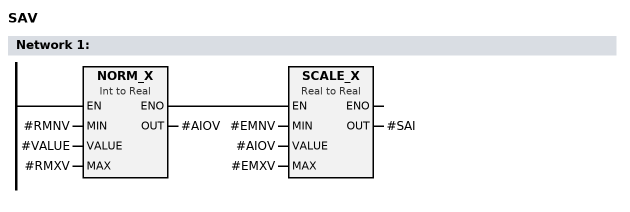
   RUNG wire#powerrail
      { S7_Templates := "[SrcType := Int, DestType := Real]" } Normalize(min := #RMNV, value := #VALUE, max := #RMXV, out => #AIOV)
      { S7_Templates := "[SrcType := Real, DestType := Real]" } Scale(min := #EMNV, value := #AIOV, max := #EMXV, out => #SAI)
   END_RUNG
   // the same network as SCL:
   #AIOV := NORM_X(MIN := #RMNV, VALUE := #VALUE, MAX := #RMXV);
   #SAI := SCALE_X(MIN := #EMNV, VALUE := #AIOV, MAX := #EMXV);
END_REGION
END_FUNCTION

// folder: 1}Library/Interlock

FUNCTION_BLOCK "Interlocks"   // FB4550, LAD
{ S7_Optimized_Access := 'TRUE' }
VERSION : 0.1
   VAR_INPUT
      Interlock_1 : Bool;
      Interlock_2 : Bool;
      Interlock_3 : Bool;
      Interlock_4 : Bool;
      Interlock_5 : Bool := false;
      Interlock_6 : Bool := false;
      Interlock_7 : Bool := false;
      Interlock_8 : Bool := false;
      Interlock_9 : Bool := false;
      Interlock_10 : Bool := false;
      Interlock_11 : Bool := false;
      Interlock_12 : Bool := false;
      Interlock_13 : Bool := false;
      Interlock_14 : Bool := false;
      Interlock_15 : Bool := false;
      Interlock_16 : Bool := false;
      Interlock_17 : Bool := false;
      Interlock_18 : Bool := false;
      Interlock_19 : Bool := false;
      Interlock_20 : Bool := false;
      Interlock_21 : Bool := false;
      Interlock_22 : Bool := false;
      Interlock_23 : Bool := false;
      Interlock_24 : Bool := false;
      Interlock_25 : Bool := false;
      Interlock_26 : Bool := false;
      Interlock_27 : Bool := false;
      Interlock_28 : Bool := false;
      Interlock_29 : Bool := false;
      Interlock_30 : Bool := false;
      Interlock_31 : Bool := false;
      Interlock_32 : Bool := false;
   END_VAR
   VAR_OUTPUT
      Out : Bool;   // Common Interlock Output
      Latched_Interlocks : DInt;   // Status of all Interlocks
   END_VAR
   VAR_IN_OUT
      Reset : Bool;
   END_VAR
   VAR
      HMI : Struct
         Interlock_1 : Bool;
         Interlock_2 : Bool;
         Interlock_3 : Bool;
         Interlock_4 : Bool;
         Interlock_5 : Bool;
         Interlock_6 : Bool;
         Interlock_7 : Bool;
         Interlock_8 : Bool;
         Interlock_9 : Bool;
         Interlock_10 : Bool;
         Interlock_11 : Bool;
         Interlock_12 : Bool;
         Interlock_13 : Bool;
         Interlock_14 : Bool;
         Interlock_15 : Bool;
         Interlock_16 : Bool;
         Interlock_17 : Bool;
         Interlock_18 : Bool;
         Interlock_19 : Bool;
         Interlock_20 : Bool;
         Interlock_21 : Bool;
         Interlock_22 : Bool;
         Interlock_23 : Bool;
         Interlock_24 : Bool;
         Interlock_25 : Bool;
         Interlock_26 : Bool;
         Interlock_27 : Bool;
         Interlock_28 : Bool;
         Interlock_29 : Bool;
         Interlock_30 : Bool;
         Interlock_31 : Bool;
         Interlock_32 : Bool;
         First_1 : Bool;
         First_2 : Bool;
         First_3 : Bool;
         First_4 : Bool;
         First_5 : Bool;
         First_6 : Bool;
         First_7 : Bool;
         First_8 : Bool;
         First_9 : Bool;
         First_10 : Bool;
         First_11 : Bool;
         First_12 : Bool;
         First_13 : Bool;
         First_14 : Bool;
         First_15 : Bool;
         First_16 : Bool;
         First_17 : Bool;
         First_18 : Bool;
         First_19 : Bool;
         First_20 : Bool;
         First_21 : Bool;
         First_22 : Bool;
         First_23 : Bool;
         First_24 : Bool;
         First_25 : Bool;
         First_26 : Bool;
         First_27 : Bool;
         First_28 : Bool;
         First_29 : Bool;
         First_30 : Bool;
         First_31 : Bool;
         First_32 : Bool;
         Bypass_1 : Bool;
         Bypass_2 : Bool;
         Bypass_3 : Bool;
         Bypass_4 : Bool;
         Bypass_5 : Bool;
         Bypass_6 : Bool;
         Bypass_7 : Bool;
         Bypass_8 : Bool;
         Bypass_9 : Bool;
         Bypass_10 : Bool;
         Bypass_11 : Bool;
         Bypass_12 : Bool;
         Bypass_13 : Bool;
         Bypass_14 : Bool;
         Bypass_15 : Bool;
         Bypass_16 : Bool;
         Bypass_17 : Bool;
         Bypass_18 : Bool;
         Bypass_19 : Bool;
         Bypass_20 : Bool;
         Bypass_21 : Bool;
         Bypass_22 : Bool;
         Bypass_23 : Bool;
         Bypass_24 : Bool;
         Bypass_25 : Bool;
         Bypass_26 : Bool;
         Bypass_27 : Bool;
         Bypass_28 : Bool;
         Bypass_29 : Bool;
         Bypass_30 : Bool;
         Bypass_31 : Bool;
         Bypass_32 : Bool;
         Status_DW : DInt;
         Interlock_DW : DInt;
         First_DW : DInt;
         Bypass_DW : DInt;
      END_STRUCT;
   END_VAR
   VAR_TEMP
      Initial_Trip : Bool;
      Interlocks_Status : DInt;
   END_VAR
BEGIN

REGION Network 1 (SCL): Common Interlock Input
   ;
   #Interlocks_Status.%X0:= #Interlock_1;
   #Interlocks_Status.%X1 := #Interlock_2;
   #Interlocks_Status.%X2 := #Interlock_3;
   #Interlocks_Status.%X3 := #Interlock_4;
   #Interlocks_Status.%X4 := #Interlock_5;
   #Interlocks_Status.%X5 := #Interlock_6;
   #Interlocks_Status.%X6 := #Interlock_7;
   #Interlocks_Status.%X7 := #Interlock_8;
   #Interlocks_Status.%X8 := #Interlock_9;
   #Interlocks_Status.%X9 := #Interlock_10;
   #Interlocks_Status.%X10 := #Interlock_11;
   #Interlocks_Status.%X11 := #Interlock_12;
   #Interlocks_Status.%X12 := #Interlock_13;
   #Interlocks_Status.%X13 := #Interlock_14;
   #Interlocks_Status.%X14 := #Interlock_15;
   #Interlocks_Status.%X15 := #Interlock_16;
   #Interlocks_Status.%X16 := #Interlock_17;
   #Interlocks_Status.%X17 := #Interlock_18;
   #Interlocks_Status.%X18 := #Interlock_19;
   #Interlocks_Status.%X19 := #Interlock_20;
   #Interlocks_Status.%X20 := #Interlock_21;
   #Interlocks_Status.%X21 := #Interlock_22;
   #Interlocks_Status.%X22 := #Interlock_23;
   #Interlocks_Status.%X23 := #Interlock_24;
   #Interlocks_Status.%X24 := #Interlock_25;
   #Interlocks_Status.%X25 := #Interlock_26;
   #Interlocks_Status.%X26 := #Interlock_27;
   #Interlocks_Status.%X27 := #Interlock_28;
   #Interlocks_Status.%X28 := #Interlock_29;
   #Interlocks_Status.%X29 := #Interlock_30;
   #Interlocks_Status.%X30 := #Interlock_31;
   #Interlocks_Status.%X31 := #Interlock_32;
END_REGION

REGION Network 2 (SCL): Bypass Move
   #HMI.Bypass_1 := #HMI.Bypass_DW.%X0;
   #HMI.Bypass_2 := #HMI.Bypass_DW.%X1;
   #HMI.Bypass_3 := #HMI.Bypass_DW.%X2;
   #HMI.Bypass_4 := #HMI.Bypass_DW.%X3;
   #HMI.Bypass_5 := #HMI.Bypass_DW.%X4;
   #HMI.Bypass_6 := #HMI.Bypass_DW.%X5;
   #HMI.Bypass_7 := #HMI.Bypass_DW.%X6;
   #HMI.Bypass_8 := #HMI.Bypass_DW.%X7;
   #HMI.Bypass_9 := #HMI.Bypass_DW.%X8;
   #HMI.Bypass_10 := #HMI.Bypass_DW.%X9;
   #HMI.Bypass_11 := #HMI.Bypass_DW.%X10;
   #HMI.Bypass_12 := #HMI.Bypass_DW.%X11;
   #HMI.Bypass_13 := #HMI.Bypass_DW.%X12;
   #HMI.Bypass_14 := #HMI.Bypass_DW.%X13;
   #HMI.Bypass_15 := #HMI.Bypass_DW.%X14;
   #HMI.Bypass_16 := #HMI.Bypass_DW.%X15;
   #HMI.Bypass_17 := #HMI.Bypass_DW.%X16;
   #HMI.Bypass_18 := #HMI.Bypass_DW.%X17;
   #HMI.Bypass_19 := #HMI.Bypass_DW.%X18;
   #HMI.Bypass_20 := #HMI.Bypass_DW.%X19;
   #HMI.Bypass_21 := #HMI.Bypass_DW.%X20;
   #HMI.Bypass_22 := #HMI.Bypass_DW.%X21;
   #HMI.Bypass_23 := #HMI.Bypass_DW.%X22;
   #HMI.Bypass_24 := #HMI.Bypass_DW.%X23;
   #HMI.Bypass_25 := #HMI.Bypass_DW.%X24;
   #HMI.Bypass_26 := #HMI.Bypass_DW.%X25;
   #HMI.Bypass_27 := #HMI.Bypass_DW.%X26;
   #HMI.Bypass_28 := #HMI.Bypass_DW.%X27;
   #HMI.Bypass_29 := #HMI.Bypass_DW.%X28;
   #HMI.Bypass_30 := #HMI.Bypass_DW.%X29;
   #HMI.Bypass_31 := #HMI.Bypass_DW.%X30;
   #HMI.Bypass_32 := #HMI.Bypass_DW.%X31;
END_REGION

REGION Network 3: Match HMI.Status_DW to Interlocks_Status
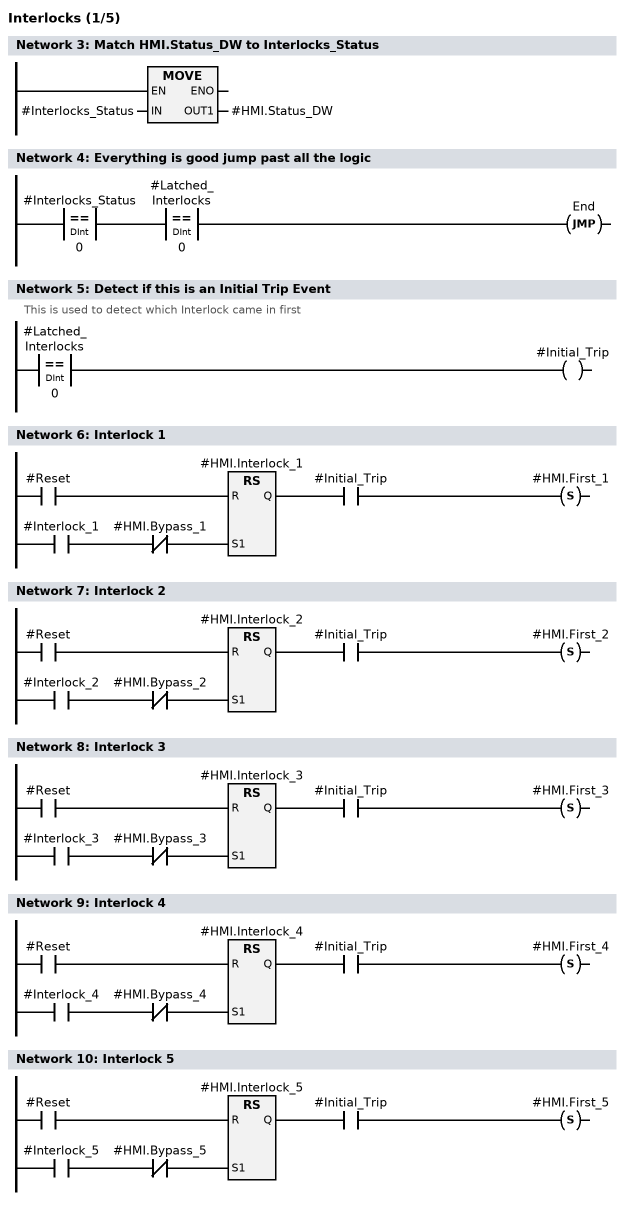
   RUNG wire#powerrail
      Move(in := #Interlocks_Status, out1 => #HMI.Status_DW)
   END_RUNG
   // the same network as SCL:
   #HMI.Status_DW := #Interlocks_Status;
END_REGION

REGION Network 4: Everything is good jump past all the logic
   RUNG wire#powerrail
      { S7_Templates := "SrcType := DInt" } EQ_Contact(in1 := #Interlocks_Status, in2 := 0)
      { S7_Templates := "SrcType := DInt" } EQ_Contact(in1 := #Latched_Interlocks, in2 := 0)
      JumpCoil( End )
   END_RUNG
   // the same network as SCL:
   IF (#Interlocks_Status = 0) AND (#Latched_Interlocks = 0) THEN GOTO End; END_IF;
END_REGION

REGION Network 5: Detect if this is an Initial Trip Event
   // This is used to detect which Interlock came in first
   RUNG wire#powerrail
      { S7_Templates := "SrcType := DInt" } EQ_Contact(in1 := #Latched_Interlocks, in2 := 0)
      Coil( #Initial_Trip )
   END_RUNG
   // the same network as SCL:
   #Initial_Trip := #Latched_Interlocks = 0;
END_REGION

REGION Network 6: Interlock 1
   RUNG wire#powerrail
      Contact( #Reset )
      S_RS(operand := #HMI.Interlock_1, s1 := wire#w1)
      Contact( #Initial_Trip )
      S_Coil( #HMI.First_1 )
   END_RUNG
   RUNG wire#powerrail
      Contact( #Interlock_1 )
      I_Contact( #HMI.Bypass_1 )
   END_RUNG wire#w1
   // the same network as SCL:
   IF #Reset THEN
       #HMI.Interlock_1 := FALSE;   // RS flip-flop
   END_IF;
   IF #Interlock_1 AND NOT #HMI.Bypass_1 THEN #HMI.Interlock_1 := TRUE; END_IF;
   IF #HMI.Interlock_1 AND #Initial_Trip THEN #HMI.First_1 := TRUE; END_IF;
END_REGION

REGION Network 7: Interlock 2
   RUNG wire#powerrail
      Contact( #Reset )
      S_RS(operand := #HMI.Interlock_2, s1 := wire#w1)
      Contact( #Initial_Trip )
      S_Coil( #HMI.First_2 )
   END_RUNG
   RUNG wire#powerrail
      Contact( #Interlock_2 )
      I_Contact( #HMI.Bypass_2 )
   END_RUNG wire#w1
   // the same network as SCL:
   IF #Reset THEN
       #HMI.Interlock_2 := FALSE;   // RS flip-flop
   END_IF;
   IF #Interlock_2 AND NOT #HMI.Bypass_2 THEN #HMI.Interlock_2 := TRUE; END_IF;
   IF #HMI.Interlock_2 AND #Initial_Trip THEN #HMI.First_2 := TRUE; END_IF;
END_REGION

REGION Network 8: Interlock 3
   RUNG wire#powerrail
      Contact( #Reset )
      S_RS(operand := #HMI.Interlock_3, s1 := wire#w1)
      Contact( #Initial_Trip )
      S_Coil( #HMI.First_3 )
   END_RUNG
   RUNG wire#powerrail
      Contact( #Interlock_3 )
      I_Contact( #HMI.Bypass_3 )
   END_RUNG wire#w1
   // the same network as SCL:
   IF #Reset THEN
       #HMI.Interlock_3 := FALSE;   // RS flip-flop
   END_IF;
   IF #Interlock_3 AND NOT #HMI.Bypass_3 THEN #HMI.Interlock_3 := TRUE; END_IF;
   IF #HMI.Interlock_3 AND #Initial_Trip THEN #HMI.First_3 := TRUE; END_IF;
END_REGION

REGION Network 9: Interlock 4
   RUNG wire#powerrail
      Contact( #Reset )
      S_RS(operand := #HMI.Interlock_4, s1 := wire#w1)
      Contact( #Initial_Trip )
      S_Coil( #HMI.First_4 )
   END_RUNG
   RUNG wire#powerrail
      Contact( #Interlock_4 )
      I_Contact( #HMI.Bypass_4 )
   END_RUNG wire#w1
   // the same network as SCL:
   IF #Reset THEN
       #HMI.Interlock_4 := FALSE;   // RS flip-flop
   END_IF;
   IF #Interlock_4 AND NOT #HMI.Bypass_4 THEN #HMI.Interlock_4 := TRUE; END_IF;
   IF #HMI.Interlock_4 AND #Initial_Trip THEN #HMI.First_4 := TRUE; END_IF;
END_REGION

REGION Network 10: Interlock 5
   RUNG wire#powerrail
      Contact( #Reset )
      S_RS(operand := #HMI.Interlock_5, s1 := wire#w1)
      Contact( #Initial_Trip )
      S_Coil( #HMI.First_5 )
   END_RUNG
   RUNG wire#powerrail
      Contact( #Interlock_5 )
      I_Contact( #HMI.Bypass_5 )
   END_RUNG wire#w1
   // the same network as SCL:
   IF #Reset THEN
       #HMI.Interlock_5 := FALSE;   // RS flip-flop
   END_IF;
   IF #Interlock_5 AND NOT #HMI.Bypass_5 THEN #HMI.Interlock_5 := TRUE; END_IF;
   IF #HMI.Interlock_5 AND #Initial_Trip THEN #HMI.First_5 := TRUE; END_IF;
END_REGION

REGION Network 11: Interlock 6
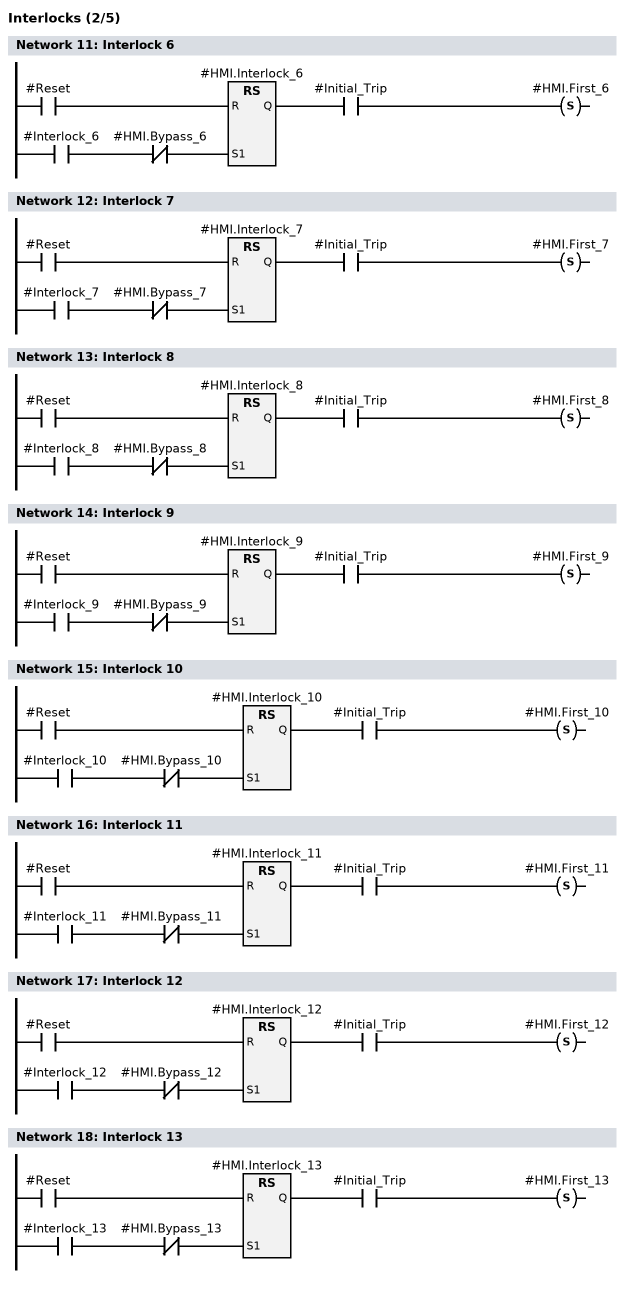
   RUNG wire#powerrail
      Contact( #Reset )
      S_RS(operand := #HMI.Interlock_6, s1 := wire#w1)
      Contact( #Initial_Trip )
      S_Coil( #HMI.First_6 )
   END_RUNG
   RUNG wire#powerrail
      Contact( #Interlock_6 )
      I_Contact( #HMI.Bypass_6 )
   END_RUNG wire#w1
   // the same network as SCL:
   IF #Reset THEN
       #HMI.Interlock_6 := FALSE;   // RS flip-flop
   END_IF;
   IF #Interlock_6 AND NOT #HMI.Bypass_6 THEN #HMI.Interlock_6 := TRUE; END_IF;
   IF #HMI.Interlock_6 AND #Initial_Trip THEN #HMI.First_6 := TRUE; END_IF;
END_REGION

REGION Network 12: Interlock 7
   RUNG wire#powerrail
      Contact( #Reset )
      S_RS(operand := #HMI.Interlock_7, s1 := wire#w1)
      Contact( #Initial_Trip )
      S_Coil( #HMI.First_7 )
   END_RUNG
   RUNG wire#powerrail
      Contact( #Interlock_7 )
      I_Contact( #HMI.Bypass_7 )
   END_RUNG wire#w1
   // the same network as SCL:
   IF #Reset THEN
       #HMI.Interlock_7 := FALSE;   // RS flip-flop
   END_IF;
   IF #Interlock_7 AND NOT #HMI.Bypass_7 THEN #HMI.Interlock_7 := TRUE; END_IF;
   IF #HMI.Interlock_7 AND #Initial_Trip THEN #HMI.First_7 := TRUE; END_IF;
END_REGION

REGION Network 13: Interlock 8
   RUNG wire#powerrail
      Contact( #Reset )
      S_RS(operand := #HMI.Interlock_8, s1 := wire#w1)
      Contact( #Initial_Trip )
      S_Coil( #HMI.First_8 )
   END_RUNG
   RUNG wire#powerrail
      Contact( #Interlock_8 )
      I_Contact( #HMI.Bypass_8 )
   END_RUNG wire#w1
   // the same network as SCL:
   IF #Reset THEN
       #HMI.Interlock_8 := FALSE;   // RS flip-flop
   END_IF;
   IF #Interlock_8 AND NOT #HMI.Bypass_8 THEN #HMI.Interlock_8 := TRUE; END_IF;
   IF #HMI.Interlock_8 AND #Initial_Trip THEN #HMI.First_8 := TRUE; END_IF;
END_REGION

REGION Network 14: Interlock 9
   RUNG wire#powerrail
      Contact( #Reset )
      S_RS(operand := #HMI.Interlock_9, s1 := wire#w1)
      Contact( #Initial_Trip )
      S_Coil( #HMI.First_9 )
   END_RUNG
   RUNG wire#powerrail
      Contact( #Interlock_9 )
      I_Contact( #HMI.Bypass_9 )
   END_RUNG wire#w1
   // the same network as SCL:
   IF #Reset THEN
       #HMI.Interlock_9 := FALSE;   // RS flip-flop
   END_IF;
   IF #Interlock_9 AND NOT #HMI.Bypass_9 THEN #HMI.Interlock_9 := TRUE; END_IF;
   IF #HMI.Interlock_9 AND #Initial_Trip THEN #HMI.First_9 := TRUE; END_IF;
END_REGION

REGION Network 15: Interlock 10
   RUNG wire#powerrail
      Contact( #Reset )
      S_RS(operand := #HMI.Interlock_10, s1 := wire#w1)
      Contact( #Initial_Trip )
      S_Coil( #HMI.First_10 )
   END_RUNG
   RUNG wire#powerrail
      Contact( #Interlock_10 )
      I_Contact( #HMI.Bypass_10 )
   END_RUNG wire#w1
   // the same network as SCL:
   IF #Reset THEN
       #HMI.Interlock_10 := FALSE;   // RS flip-flop
   END_IF;
   IF #Interlock_10 AND NOT #HMI.Bypass_10 THEN #HMI.Interlock_10 := TRUE; END_IF;
   IF #HMI.Interlock_10 AND #Initial_Trip THEN #HMI.First_10 := TRUE; END_IF;
END_REGION

REGION Network 16: Interlock 11
   RUNG wire#powerrail
      Contact( #Reset )
      S_RS(operand := #HMI.Interlock_11, s1 := wire#w1)
      Contact( #Initial_Trip )
      S_Coil( #HMI.First_11 )
   END_RUNG
   RUNG wire#powerrail
      Contact( #Interlock_11 )
      I_Contact( #HMI.Bypass_11 )
   END_RUNG wire#w1
   // the same network as SCL:
   IF #Reset THEN
       #HMI.Interlock_11 := FALSE;   // RS flip-flop
   END_IF;
   IF #Interlock_11 AND NOT #HMI.Bypass_11 THEN #HMI.Interlock_11 := TRUE; END_IF;
   IF #HMI.Interlock_11 AND #Initial_Trip THEN #HMI.First_11 := TRUE; END_IF;
END_REGION

REGION Network 17: Interlock 12
   RUNG wire#powerrail
      Contact( #Reset )
      S_RS(operand := #HMI.Interlock_12, s1 := wire#w1)
      Contact( #Initial_Trip )
      S_Coil( #HMI.First_12 )
   END_RUNG
   RUNG wire#powerrail
      Contact( #Interlock_12 )
      I_Contact( #HMI.Bypass_12 )
   END_RUNG wire#w1
   // the same network as SCL:
   IF #Reset THEN
       #HMI.Interlock_12 := FALSE;   // RS flip-flop
   END_IF;
   IF #Interlock_12 AND NOT #HMI.Bypass_12 THEN #HMI.Interlock_12 := TRUE; END_IF;
   IF #HMI.Interlock_12 AND #Initial_Trip THEN #HMI.First_12 := TRUE; END_IF;
END_REGION

REGION Network 18: Interlock 13
   RUNG wire#powerrail
      Contact( #Reset )
      S_RS(operand := #HMI.Interlock_13, s1 := wire#w1)
      Contact( #Initial_Trip )
      S_Coil( #HMI.First_13 )
   END_RUNG
   RUNG wire#powerrail
      Contact( #Interlock_13 )
      I_Contact( #HMI.Bypass_13 )
   END_RUNG wire#w1
   // the same network as SCL:
   IF #Reset THEN
       #HMI.Interlock_13 := FALSE;   // RS flip-flop
   END_IF;
   IF #Interlock_13 AND NOT #HMI.Bypass_13 THEN #HMI.Interlock_13 := TRUE; END_IF;
   IF #HMI.Interlock_13 AND #Initial_Trip THEN #HMI.First_13 := TRUE; END_IF;
END_REGION

REGION Network 19: Interlock 14
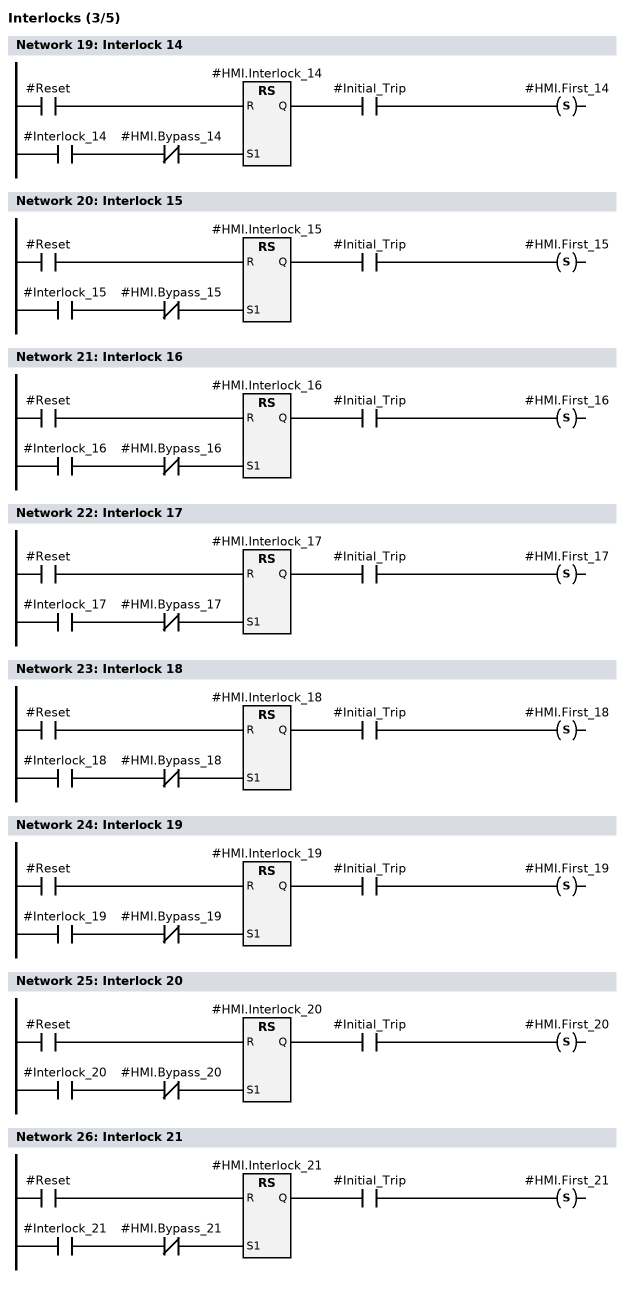
   RUNG wire#powerrail
      Contact( #Reset )
      S_RS(operand := #HMI.Interlock_14, s1 := wire#w1)
      Contact( #Initial_Trip )
      S_Coil( #HMI.First_14 )
   END_RUNG
   RUNG wire#powerrail
      Contact( #Interlock_14 )
      I_Contact( #HMI.Bypass_14 )
   END_RUNG wire#w1
   // the same network as SCL:
   IF #Reset THEN
       #HMI.Interlock_14 := FALSE;   // RS flip-flop
   END_IF;
   IF #Interlock_14 AND NOT #HMI.Bypass_14 THEN #HMI.Interlock_14 := TRUE; END_IF;
   IF #HMI.Interlock_14 AND #Initial_Trip THEN #HMI.First_14 := TRUE; END_IF;
END_REGION

REGION Network 20: Interlock 15
   RUNG wire#powerrail
      Contact( #Reset )
      S_RS(operand := #HMI.Interlock_15, s1 := wire#w1)
      Contact( #Initial_Trip )
      S_Coil( #HMI.First_15 )
   END_RUNG
   RUNG wire#powerrail
      Contact( #Interlock_15 )
      I_Contact( #HMI.Bypass_15 )
   END_RUNG wire#w1
   // the same network as SCL:
   IF #Reset THEN
       #HMI.Interlock_15 := FALSE;   // RS flip-flop
   END_IF;
   IF #Interlock_15 AND NOT #HMI.Bypass_15 THEN #HMI.Interlock_15 := TRUE; END_IF;
   IF #HMI.Interlock_15 AND #Initial_Trip THEN #HMI.First_15 := TRUE; END_IF;
END_REGION

REGION Network 21: Interlock 16
   RUNG wire#powerrail
      Contact( #Reset )
      S_RS(operand := #HMI.Interlock_16, s1 := wire#w1)
      Contact( #Initial_Trip )
      S_Coil( #HMI.First_16 )
   END_RUNG
   RUNG wire#powerrail
      Contact( #Interlock_16 )
      I_Contact( #HMI.Bypass_16 )
   END_RUNG wire#w1
   // the same network as SCL:
   IF #Reset THEN
       #HMI.Interlock_16 := FALSE;   // RS flip-flop
   END_IF;
   IF #Interlock_16 AND NOT #HMI.Bypass_16 THEN #HMI.Interlock_16 := TRUE; END_IF;
   IF #HMI.Interlock_16 AND #Initial_Trip THEN #HMI.First_16 := TRUE; END_IF;
END_REGION

REGION Network 22: Interlock 17
   RUNG wire#powerrail
      Contact( #Reset )
      S_RS(operand := #HMI.Interlock_17, s1 := wire#w1)
      Contact( #Initial_Trip )
      S_Coil( #HMI.First_17 )
   END_RUNG
   RUNG wire#powerrail
      Contact( #Interlock_17 )
      I_Contact( #HMI.Bypass_17 )
   END_RUNG wire#w1
   // the same network as SCL:
   IF #Reset THEN
       #HMI.Interlock_17 := FALSE;   // RS flip-flop
   END_IF;
   IF #Interlock_17 AND NOT #HMI.Bypass_17 THEN #HMI.Interlock_17 := TRUE; END_IF;
   IF #HMI.Interlock_17 AND #Initial_Trip THEN #HMI.First_17 := TRUE; END_IF;
END_REGION

REGION Network 23: Interlock 18
   RUNG wire#powerrail
      Contact( #Reset )
      S_RS(operand := #HMI.Interlock_18, s1 := wire#w1)
      Contact( #Initial_Trip )
      S_Coil( #HMI.First_18 )
   END_RUNG
   RUNG wire#powerrail
      Contact( #Interlock_18 )
      I_Contact( #HMI.Bypass_18 )
   END_RUNG wire#w1
   // the same network as SCL:
   IF #Reset THEN
       #HMI.Interlock_18 := FALSE;   // RS flip-flop
   END_IF;
   IF #Interlock_18 AND NOT #HMI.Bypass_18 THEN #HMI.Interlock_18 := TRUE; END_IF;
   IF #HMI.Interlock_18 AND #Initial_Trip THEN #HMI.First_18 := TRUE; END_IF;
END_REGION

REGION Network 24: Interlock 19
   RUNG wire#powerrail
      Contact( #Reset )
      S_RS(operand := #HMI.Interlock_19, s1 := wire#w1)
      Contact( #Initial_Trip )
      S_Coil( #HMI.First_19 )
   END_RUNG
   RUNG wire#powerrail
      Contact( #Interlock_19 )
      I_Contact( #HMI.Bypass_19 )
   END_RUNG wire#w1
   // the same network as SCL:
   IF #Reset THEN
       #HMI.Interlock_19 := FALSE;   // RS flip-flop
   END_IF;
   IF #Interlock_19 AND NOT #HMI.Bypass_19 THEN #HMI.Interlock_19 := TRUE; END_IF;
   IF #HMI.Interlock_19 AND #Initial_Trip THEN #HMI.First_19 := TRUE; END_IF;
END_REGION

REGION Network 25: Interlock 20
   RUNG wire#powerrail
      Contact( #Reset )
      S_RS(operand := #HMI.Interlock_20, s1 := wire#w1)
      Contact( #Initial_Trip )
      S_Coil( #HMI.First_20 )
   END_RUNG
   RUNG wire#powerrail
      Contact( #Interlock_20 )
      I_Contact( #HMI.Bypass_20 )
   END_RUNG wire#w1
   // the same network as SCL:
   IF #Reset THEN
       #HMI.Interlock_20 := FALSE;   // RS flip-flop
   END_IF;
   IF #Interlock_20 AND NOT #HMI.Bypass_20 THEN #HMI.Interlock_20 := TRUE; END_IF;
   IF #HMI.Interlock_20 AND #Initial_Trip THEN #HMI.First_20 := TRUE; END_IF;
END_REGION

REGION Network 26: Interlock 21
   RUNG wire#powerrail
      Contact( #Reset )
      S_RS(operand := #HMI.Interlock_21, s1 := wire#w1)
      Contact( #Initial_Trip )
      S_Coil( #HMI.First_21 )
   END_RUNG
   RUNG wire#powerrail
      Contact( #Interlock_21 )
      I_Contact( #HMI.Bypass_21 )
   END_RUNG wire#w1
   // the same network as SCL:
   IF #Reset THEN
       #HMI.Interlock_21 := FALSE;   // RS flip-flop
   END_IF;
   IF #Interlock_21 AND NOT #HMI.Bypass_21 THEN #HMI.Interlock_21 := TRUE; END_IF;
   IF #HMI.Interlock_21 AND #Initial_Trip THEN #HMI.First_21 := TRUE; END_IF;
END_REGION

REGION Network 27: Interlock 22
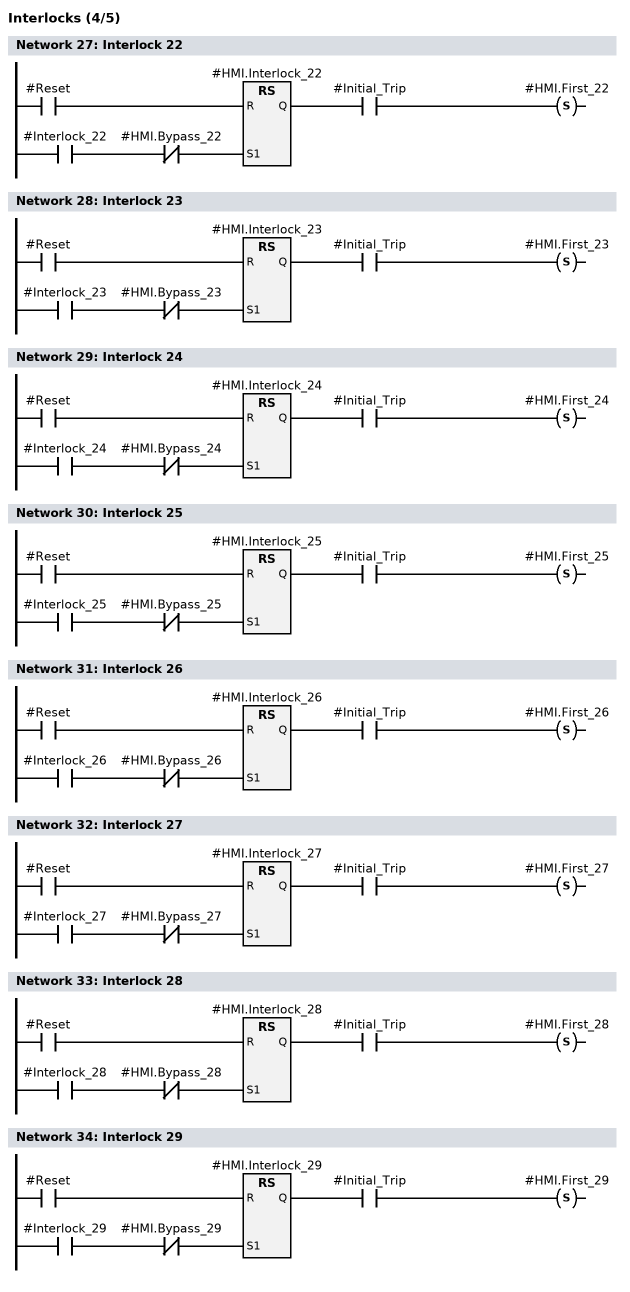
   RUNG wire#powerrail
      Contact( #Reset )
      S_RS(operand := #HMI.Interlock_22, s1 := wire#w1)
      Contact( #Initial_Trip )
      S_Coil( #HMI.First_22 )
   END_RUNG
   RUNG wire#powerrail
      Contact( #Interlock_22 )
      I_Contact( #HMI.Bypass_22 )
   END_RUNG wire#w1
   // the same network as SCL:
   IF #Reset THEN
       #HMI.Interlock_22 := FALSE;   // RS flip-flop
   END_IF;
   IF #Interlock_22 AND NOT #HMI.Bypass_22 THEN #HMI.Interlock_22 := TRUE; END_IF;
   IF #HMI.Interlock_22 AND #Initial_Trip THEN #HMI.First_22 := TRUE; END_IF;
END_REGION

REGION Network 28: Interlock 23
   RUNG wire#powerrail
      Contact( #Reset )
      S_RS(operand := #HMI.Interlock_23, s1 := wire#w1)
      Contact( #Initial_Trip )
      S_Coil( #HMI.First_23 )
   END_RUNG
   RUNG wire#powerrail
      Contact( #Interlock_23 )
      I_Contact( #HMI.Bypass_23 )
   END_RUNG wire#w1
   // the same network as SCL:
   IF #Reset THEN
       #HMI.Interlock_23 := FALSE;   // RS flip-flop
   END_IF;
   IF #Interlock_23 AND NOT #HMI.Bypass_23 THEN #HMI.Interlock_23 := TRUE; END_IF;
   IF #HMI.Interlock_23 AND #Initial_Trip THEN #HMI.First_23 := TRUE; END_IF;
END_REGION

REGION Network 29: Interlock 24
   RUNG wire#powerrail
      Contact( #Reset )
      S_RS(operand := #HMI.Interlock_24, s1 := wire#w1)
      Contact( #Initial_Trip )
      S_Coil( #HMI.First_24 )
   END_RUNG
   RUNG wire#powerrail
      Contact( #Interlock_24 )
      I_Contact( #HMI.Bypass_24 )
   END_RUNG wire#w1
   // the same network as SCL:
   IF #Reset THEN
       #HMI.Interlock_24 := FALSE;   // RS flip-flop
   END_IF;
   IF #Interlock_24 AND NOT #HMI.Bypass_24 THEN #HMI.Interlock_24 := TRUE; END_IF;
   IF #HMI.Interlock_24 AND #Initial_Trip THEN #HMI.First_24 := TRUE; END_IF;
END_REGION

REGION Network 30: Interlock 25
   RUNG wire#powerrail
      Contact( #Reset )
      S_RS(operand := #HMI.Interlock_25, s1 := wire#w1)
      Contact( #Initial_Trip )
      S_Coil( #HMI.First_25 )
   END_RUNG
   RUNG wire#powerrail
      Contact( #Interlock_25 )
      I_Contact( #HMI.Bypass_25 )
   END_RUNG wire#w1
   // the same network as SCL:
   IF #Reset THEN
       #HMI.Interlock_25 := FALSE;   // RS flip-flop
   END_IF;
   IF #Interlock_25 AND NOT #HMI.Bypass_25 THEN #HMI.Interlock_25 := TRUE; END_IF;
   IF #HMI.Interlock_25 AND #Initial_Trip THEN #HMI.First_25 := TRUE; END_IF;
END_REGION

REGION Network 31: Interlock 26
   RUNG wire#powerrail
      Contact( #Reset )
      S_RS(operand := #HMI.Interlock_26, s1 := wire#w1)
      Contact( #Initial_Trip )
      S_Coil( #HMI.First_26 )
   END_RUNG
   RUNG wire#powerrail
      Contact( #Interlock_26 )
      I_Contact( #HMI.Bypass_26 )
   END_RUNG wire#w1
   // the same network as SCL:
   IF #Reset THEN
       #HMI.Interlock_26 := FALSE;   // RS flip-flop
   END_IF;
   IF #Interlock_26 AND NOT #HMI.Bypass_26 THEN #HMI.Interlock_26 := TRUE; END_IF;
   IF #HMI.Interlock_26 AND #Initial_Trip THEN #HMI.First_26 := TRUE; END_IF;
END_REGION

REGION Network 32: Interlock 27
   RUNG wire#powerrail
      Contact( #Reset )
      S_RS(operand := #HMI.Interlock_27, s1 := wire#w1)
      Contact( #Initial_Trip )
      S_Coil( #HMI.First_27 )
   END_RUNG
   RUNG wire#powerrail
      Contact( #Interlock_27 )
      I_Contact( #HMI.Bypass_27 )
   END_RUNG wire#w1
   // the same network as SCL:
   IF #Reset THEN
       #HMI.Interlock_27 := FALSE;   // RS flip-flop
   END_IF;
   IF #Interlock_27 AND NOT #HMI.Bypass_27 THEN #HMI.Interlock_27 := TRUE; END_IF;
   IF #HMI.Interlock_27 AND #Initial_Trip THEN #HMI.First_27 := TRUE; END_IF;
END_REGION

REGION Network 33: Interlock 28
   RUNG wire#powerrail
      Contact( #Reset )
      S_RS(operand := #HMI.Interlock_28, s1 := wire#w1)
      Contact( #Initial_Trip )
      S_Coil( #HMI.First_28 )
   END_RUNG
   RUNG wire#powerrail
      Contact( #Interlock_28 )
      I_Contact( #HMI.Bypass_28 )
   END_RUNG wire#w1
   // the same network as SCL:
   IF #Reset THEN
       #HMI.Interlock_28 := FALSE;   // RS flip-flop
   END_IF;
   IF #Interlock_28 AND NOT #HMI.Bypass_28 THEN #HMI.Interlock_28 := TRUE; END_IF;
   IF #HMI.Interlock_28 AND #Initial_Trip THEN #HMI.First_28 := TRUE; END_IF;
END_REGION

REGION Network 34: Interlock 29
   RUNG wire#powerrail
      Contact( #Reset )
      S_RS(operand := #HMI.Interlock_29, s1 := wire#w1)
      Contact( #Initial_Trip )
      S_Coil( #HMI.First_29 )
   END_RUNG
   RUNG wire#powerrail
      Contact( #Interlock_29 )
      I_Contact( #HMI.Bypass_29 )
   END_RUNG wire#w1
   // the same network as SCL:
   IF #Reset THEN
       #HMI.Interlock_29 := FALSE;   // RS flip-flop
   END_IF;
   IF #Interlock_29 AND NOT #HMI.Bypass_29 THEN #HMI.Interlock_29 := TRUE; END_IF;
   IF #HMI.Interlock_29 AND #Initial_Trip THEN #HMI.First_29 := TRUE; END_IF;
END_REGION

REGION Network 35: Interlock 30
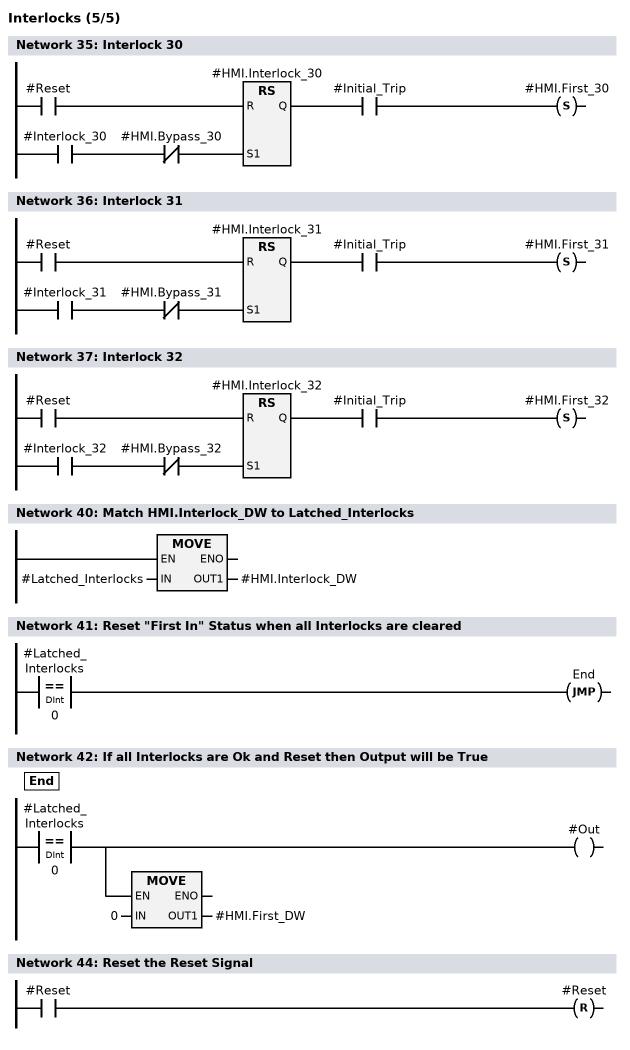
   RUNG wire#powerrail
      Contact( #Reset )
      S_RS(operand := #HMI.Interlock_30, s1 := wire#w1)
      Contact( #Initial_Trip )
      S_Coil( #HMI.First_30 )
   END_RUNG
   RUNG wire#powerrail
      Contact( #Interlock_30 )
      I_Contact( #HMI.Bypass_30 )
   END_RUNG wire#w1
   // the same network as SCL:
   IF #Reset THEN
       #HMI.Interlock_30 := FALSE;   // RS flip-flop
   END_IF;
   IF #Interlock_30 AND NOT #HMI.Bypass_30 THEN #HMI.Interlock_30 := TRUE; END_IF;
   IF #HMI.Interlock_30 AND #Initial_Trip THEN #HMI.First_30 := TRUE; END_IF;
END_REGION

REGION Network 36: Interlock 31
   RUNG wire#powerrail
      Contact( #Reset )
      S_RS(operand := #HMI.Interlock_31, s1 := wire#w1)
      Contact( #Initial_Trip )
      S_Coil( #HMI.First_31 )
   END_RUNG
   RUNG wire#powerrail
      Contact( #Interlock_31 )
      I_Contact( #HMI.Bypass_31 )
   END_RUNG wire#w1
   // the same network as SCL:
   IF #Reset THEN
       #HMI.Interlock_31 := FALSE;   // RS flip-flop
   END_IF;
   IF #Interlock_31 AND NOT #HMI.Bypass_31 THEN #HMI.Interlock_31 := TRUE; END_IF;
   IF #HMI.Interlock_31 AND #Initial_Trip THEN #HMI.First_31 := TRUE; END_IF;
END_REGION

REGION Network 37: Interlock 32
   RUNG wire#powerrail
      Contact( #Reset )
      S_RS(operand := #HMI.Interlock_32, s1 := wire#w1)
      Contact( #Initial_Trip )
      S_Coil( #HMI.First_32 )
   END_RUNG
   RUNG wire#powerrail
      Contact( #Interlock_32 )
      I_Contact( #HMI.Bypass_32 )
   END_RUNG wire#w1
   // the same network as SCL:
   IF #Reset THEN
       #HMI.Interlock_32 := FALSE;   // RS flip-flop
   END_IF;
   IF #Interlock_32 AND NOT #HMI.Bypass_32 THEN #HMI.Interlock_32 := TRUE; END_IF;
   IF #HMI.Interlock_32 AND #Initial_Trip THEN #HMI.First_32 := TRUE; END_IF;
END_REGION

REGION Network 38 (SCL): First In
   #HMI.First_DW.%X0 := #HMI.First_1;
   #HMI.First_DW.%X1 := #HMI.First_2;
   #HMI.First_DW.%X2 := #HMI.First_3;
   #HMI.First_DW.%X3 := #HMI.First_4;
   #HMI.First_DW.%X4 := #HMI.First_5;
   #HMI.First_DW.%X5 := #HMI.First_6;
   #HMI.First_DW.%X6 := #HMI.First_7;
   #HMI.First_DW.%X7 := #HMI.First_8;
   #HMI.First_DW.%X8 := #HMI.First_9;
   #HMI.First_DW.%X9 := #HMI.First_10;
   #HMI.First_DW.%X10 := #HMI.First_11;
   #HMI.First_DW.%X11 := #HMI.First_12;
   #HMI.First_DW.%X12 := #HMI.First_13;
   #HMI.First_DW.%X13 := #HMI.First_14;
   #HMI.First_DW.%X14 := #HMI.First_15;
   #HMI.First_DW.%X15 := #HMI.First_16;
   #HMI.First_DW.%X16 := #HMI.First_17;
   #HMI.First_DW.%X17 := #HMI.First_18;
   #HMI.First_DW.%X18 := #HMI.First_19;
   #HMI.First_DW.%X19 := #HMI.First_20;
   #HMI.First_DW.%X20 := #HMI.First_21;
   #HMI.First_DW.%X21 := #HMI.First_22;
   #HMI.First_DW.%X22 := #HMI.First_23;
   #HMI.First_DW.%X23 := #HMI.First_24;
   #HMI.First_DW.%X24 := #HMI.First_25;
   #HMI.First_DW.%X25 := #HMI.First_26;
   #HMI.First_DW.%X26 := #HMI.First_27;
   #HMI.First_DW.%X27 := #HMI.First_28;
   #HMI.First_DW.%X28 := #HMI.First_29;
   #HMI.First_DW.%X29 := #HMI.First_30;
   #HMI.First_DW.%X30 := #HMI.First_31;
   #HMI.First_DW.%X31 := #HMI.First_32;
END_REGION

REGION Network 39 (SCL): Common Interlock Output
   ;
   #Latched_Interlocks.%X0:= #HMI.Interlock_1;
   #Latched_Interlocks.%X1 := #HMI.Interlock_2;
   #Latched_Interlocks.%X2 := #HMI.Interlock_3;
   #Latched_Interlocks.%X3 := #HMI.Interlock_4;
   #Latched_Interlocks.%X4 := #HMI.Interlock_5;
   #Latched_Interlocks.%X5 := #HMI.Interlock_6;
   #Latched_Interlocks.%X6 := #HMI.Interlock_7;
   #Latched_Interlocks.%X7 := #HMI.Interlock_8;
   #Latched_Interlocks.%X8 := #HMI.Interlock_9;
   #Latched_Interlocks.%X9 := #HMI.Interlock_10;
   #Latched_Interlocks.%X10 := #HMI.Interlock_11;
   #Latched_Interlocks.%X11 := #HMI.Interlock_12;
   #Latched_Interlocks.%X12 := #HMI.Interlock_13;
   #Latched_Interlocks.%X13 := #HMI.Interlock_14;
   #Latched_Interlocks.%X14 := #HMI.Interlock_15;
   #Latched_Interlocks.%X15 := #HMI.Interlock_16;
   #Latched_Interlocks.%X16 := #HMI.Interlock_17;
   #Latched_Interlocks.%X17 := #HMI.Interlock_18;
   #Latched_Interlocks.%X18 := #HMI.Interlock_19;
   #Latched_Interlocks.%X19 := #HMI.Interlock_20;
   #Latched_Interlocks.%X20 := #HMI.Interlock_21;
   #Latched_Interlocks.%X21 := #HMI.Interlock_22;
   #Latched_Interlocks.%X22 := #HMI.Interlock_23;
   #Latched_Interlocks.%X23 := #HMI.Interlock_24;
   #Latched_Interlocks.%X24 := #HMI.Interlock_25;
   #Latched_Interlocks.%X25 := #HMI.Interlock_26;
   #Latched_Interlocks.%X26 := #HMI.Interlock_27;
   #Latched_Interlocks.%X27 := #HMI.Interlock_28;
   #Latched_Interlocks.%X28 := #HMI.Interlock_29;
   #Latched_Interlocks.%X29 := #HMI.Interlock_30;
   #Latched_Interlocks.%X30 := #HMI.Interlock_31;
   #Latched_Interlocks.%X31 := #HMI.Interlock_32;
END_REGION

REGION Network 40: Match HMI.Interlock_DW to Latched_Interlocks
   RUNG wire#powerrail
      Move(in := #Latched_Interlocks, out1 => #HMI.Interlock_DW)
   END_RUNG
   // the same network as SCL:
   #HMI.Interlock_DW := #Latched_Interlocks;
END_REGION

REGION Network 41: Reset "First In" Status when all Interlocks are cleared
   RUNG wire#powerrail
      { S7_Templates := "SrcType := DInt" } EQ_Contact(in1 := #Latched_Interlocks, in2 := 0)
      JumpCoil( End )
   END_RUNG
   // the same network as SCL:
   IF #Latched_Interlocks = 0 THEN GOTO End; END_IF;
END_REGION

REGION Network 42: If all Interlocks are Ok and Reset then Output will be True
   Label( End )
   RUNG wire#powerrail
      { S7_Templates := "SrcType := DInt" } EQ_Contact(in1 := #Latched_Interlocks, in2 := 0)
      wire#w1
      Coil( #Out )
   END_RUNG
   RUNG wire#w1
      { S7_GenerateENO := "TRUE" } Move(in := 0, out1 => #HMI.First_DW)
   END_RUNG
   // the same network as SCL:
   End:
   #Out := #Latched_Interlocks = 0;
   IF #Out THEN #HMI.First_DW := 0; END_IF;
END_REGION

REGION Network 43 (SCL)
   IF #Latched_Interlocks = 0 THEN
       #HMI.First_1 := 0;
       #HMI.First_2 := 0;
       #HMI.First_3 := 0;
       #HMI.First_4 := 0;
       #HMI.First_5 := 0;
       #HMI.First_6 := 0;
       #HMI.First_7 := 0;
       #HMI.First_8 := 0;
       #HMI.First_9 := 0;
       #HMI.First_10 := 0;
       #HMI.First_11 := 0;
       #HMI.First_12 := 0;
       #HMI.First_13 := 0;
       #HMI.First_14 := 0;
       #HMI.First_15 := 0;
       #HMI.First_16 := 0;
       #HMI.First_17 := 0;
       #HMI.First_18 := 0;
       #HMI.First_19 := 0;
       #HMI.First_20 := 0;
       #HMI.First_21 := 0;
       #HMI.First_22 := 0;
       #HMI.First_23 := 0;
       #HMI.First_24 := 0;
       #HMI.First_25 := 0;
       #HMI.First_26 := 0;
       #HMI.First_27 := 0;
       #HMI.First_28 := 0;
       #HMI.First_29 := 0;
       #HMI.First_30 := 0;
       #HMI.First_31 := 0;
       #HMI.First_32 := 0;
   END_IF;
END_REGION

REGION Network 44: Reset the Reset Signal
   RUNG wire#powerrail
      Contact( #Reset )
      R_Coil( #Reset )
   END_RUNG
   // the same network as SCL:
   IF #Reset THEN #Reset := FALSE; END_IF;
END_REGION
END_FUNCTION_BLOCK

// folder: 1}Library/MotorStarterET200SP

FUNCTION_BLOCK "MotorStarterET200SPchanged"   // FB813, LAD
{ S7_Optimized_Access := 'TRUE' }